// TIA Portal project "Parsing_migrated" (V16) (continued)
TYPE "LKinLang_typeKeyToken"
   STRUCT
      tokenBool : String["LKINLANG_LENGTH_OF_TOKEN_STRING"] := 'BOOL';   // Keyword for dataType "BOOL"
      tokenDInt : String["LKINLANG_LENGTH_OF_TOKEN_STRING"] := 'DINT';   // Keyword for dataType "DINT"
      tokenLReal : String["LKINLANG_LENGTH_OF_TOKEN_STRING"] := 'LREAL';   // Keyword for dataType "LREAL"
      tokenInterfaceVarBool : String["LKINLANG_LENGTH_OF_TOKEN_STRING"] := '%B';   // Keyword for interface variable type "BOOL"
      tokenInterfaceVarDInt : String["LKINLANG_LENGTH_OF_TOKEN_STRING"] := '%DI';   // Keyword for interface variable type "DINT"
      tokenInterfaceVarLReal : String["LKINLANG_LENGTH_OF_TOKEN_STRING"] := '%LR';   // Keyword for interface variable type "LREAL"
      tokenJumpTarget : String["LKINLANG_LENGTH_OF_TOKEN_STRING"] := 'LABEL';   // Keyword for label definition
      tokenJump : String["LKINLANG_LENGTH_OF_TOKEN_STRING"] := 'GOTO';   // Keyword for unconditional jump
      tokenJumpConditional : String["LKINLANG_LENGTH_OF_TOKEN_STRING"] := 'GOTOC';   // Keyword for conditional jump
      tokenPreprocessingStop : String["LKINLANG_LENGTH_OF_TOKEN_STRING"] := 'STOPRE';   // Keyword for preprocessing stop
      tokenIf : String["LKINLANG_LENGTH_OF_TOKEN_STRING"] := 'IF';   // Keyword for start of IF
      tokenElse : String["LKINLANG_LENGTH_OF_TOKEN_STRING"] := 'ELSE';   // Keyword for ELSE / Keyword for Else
      tokenEndIf : String["LKINLANG_LENGTH_OF_TOKEN_STRING"] := 'ENDIF';   // Keyword for end of IF / Keyword for end of if
      tokenWhile : String["LKINLANG_LENGTH_OF_TOKEN_STRING"] := 'WHILE';   // Keyword for start of WHILE
      tokenEndWhile : String["LKINLANG_LENGTH_OF_TOKEN_STRING"] := 'ENDWHILE';   // Keyword for end of WHILE
      tokenFor : String["LKINLANG_LENGTH_OF_TOKEN_STRING"] := 'FOR';   // Keyword for start of FOR
      tokenQuantity : String["LKINLANG_LENGTH_OF_TOKEN_STRING"] := 'TO';   // Keyword for end value of FOR
      tokenIncrement : String["LKINLANG_LENGTH_OF_TOKEN_STRING"] := 'STEP';   // Keyword for increment of FOR
      tokenEndFor : String["LKINLANG_LENGTH_OF_TOKEN_STRING"] := 'ENDFOR';   // Keyword for end of FOR
      tokenStartSub : String["LKINLANG_LENGTH_OF_TOKEN_STRING"] := 'SUB';   // Keyword for starting the definition of a subprogram
      tokenEndSub : String["LKINLANG_LENGTH_OF_TOKEN_STRING"] := 'ENDSUB';   // Keyword for ending the definition of a subprogram
      tokenCallSub : String["LKINLANG_LENGTH_OF_TOKEN_STRING"] := 'CALL';   // Keyword for calling a subprogram
      tokenReturnSub : String["LKINLANG_LENGTH_OF_TOKEN_STRING"] := 'RETURN';   // Keyword for returning from a subprogram
   END_STRUCT;
END_TYPE

TYPE "LKinLang_typeFlagModeDefaults"
   STRUCT
      setFlags : Array[0.."LKINCTRL_NO_OF_LAST_SETFLAG"] of "LKinLang_typeFlagModeDefaultElement";   // Default flag settings for respective setFlag number
      valueFlags : Array[0.."LKINCTRL_NO_OF_LAST_VALUEFLAG"] of "LKinLang_typeFlagModeDefaultElement";   // Default flag settings for respective valueFlag number
   END_STRUCT;
END_TYPE

TYPE "LKinLang_typeLineTokens"
   STRUCT
      lineNo : UDInt;   // line number
      numberOfToken : DInt;   // number of token
      lineToken : Array[1.."LKINLANG_MAX_NUMBER_OF_TOKEN_PER_LINE"] of String["LKINLANG_LENGTH_OF_TOKEN_STRING"];   // array of line tokens
   END_STRUCT;
END_TYPE

TYPE "LKinLang_typeMathParserResult"
   STRUCT
      finalResult : LReal;   // final result of math parser
      errorID : DInt;   // error code of math parser calculation
   END_STRUCT;
END_TYPE

TYPE "LKinLang_typeDiffElementaryDatatypes"
   STRUCT
      valueLReal : LReal;   // LReal value
      valueReal : Real;   // Real value
      valueDint : DInt;   // DInt value
      valueInt : Int;   // Int value
   END_STRUCT;
END_TYPE

TYPE "LKinLang_typeFlagModeDefaultElement"
   STRUCT
      flagMode : USInt;   // Default flag mode for respective setFlag number
      remainingDistance : LReal;   // Default remainingDistance for respective setFlag number in case of flagMode = 10
   END_STRUCT;
END_TYPE

TYPE "LKinLang_typePreProcessorReplacement"
   STRUCT
      replacements : Array[1.."LKINLANG_NUMBER_OF_REPLACEMENTS"] of Struct   // pre-processor replacement structure
         searchTerm : String["LKINLANG_MAX_NUMBER_OF_TOKEN_PER_LINE"];   // term to be searched
         replaceTerm : String["LKINLANG_MAX_NUMBER_OF_TOKEN_PER_LINE"];   // term to replace search term
      END_STRUCT;
   END_STRUCT;
END_TYPE

TYPE "LKinLang_typeGCodeDefaults"
   STRUCT
      velocityRapidLinear : LReal := -1.0;   // velocity for G0 command / velocity for FastLin command
      transitionVelocityMode : DInt := 5;   // Set G641 transition velocity (bufferMode); 2: low velocity, 5: high velocity
      orientationDirection : DInt := 3;   // Set orientation direction; 1: positive direction; 2: negative direction; 3: shortest distance
   END_STRUCT;
END_TYPE

TYPE "LKInLang_typeStackElement"
   STRUCT
      "type" : Int;   // Type of stack entry
      lineNumberStart : UDInt;   // Line number where stack entry starts
      lineNumberEnd : UDInt;   // Line number where stack entry ends
      variableRef : "LKinLang_typeVarRef";   // Counter variable reference (only for FOR loops)
      increment : DInt;   // Increment of FOR loop
      quantity : DInt;   // End value of FOR loop
   END_STRUCT;
END_TYPE

TYPE "LKInLang_typeHierarchicLevel"
   STRUCT
      currentLevel : Int;   // Current hierarchic level
      numberOfLevels : Int;   // Number of found hierarchic level changes
      levels : Array[1.."LKINLANG_NUMBER_OF_HIERARCHICLEVEL"] of "LKInLang_typeHierarchicLevelElement";   // Array of level changes
   END_STRUCT;
END_TYPE

TYPE "LKinLang_typeStack"
   STRUCT
      numberOfElements : Int;   // Counter for stack elements
      stackElements : Array[1..20] of "LKInLang_typeStackElement";   // Array of stack entries
   END_STRUCT;
END_TYPE

TYPE "LKInLang_typeHierarchicLevelElement"
   STRUCT
      lineNumber : UDInt;   // Line number where new hierarchic level start
      level : Int;   // Value of hierarchic level
      "type" : Int;   // Type of hierarchic level
   END_STRUCT;
END_TYPE

TYPE "LKinLang_typeSubPrg"
   STRUCT
      prgName : String;   // Name of subprogram
      lineNumberStart : UDInt;   // Line number where subprograms starts
      lineNumberEnd : UDInt;   // Line number where subprograms ends
   END_STRUCT;
END_TYPE

TYPE "LKinLang_typeSubPrgList"
   STRUCT
      numberOfSubPrgs : Int;   // Counter of found subprograms
      subPrgs : Array[1.."LKINLANG_NUMBER_OF_SUBPROGRAMS"] of "LKinLang_typeSubPrg";   // Array of subprograms
   END_STRUCT;
END_TYPE

TYPE "LKinLang_typeVariableDeclaration"
   STRUCT
      localVariables : String := 'DEF _type_ _name_';   // How to declare a local variable
      globalVariables : String := 'DEF GLOBAL _type_ _name_';   // How to declare a global variable
   END_STRUCT;
END_TYPE

TYPE "LKinLang_typeParameterDefinition"
   STRUCT
      parameterNameString : String;   // parameter name (textual)
      parameterNameNumber : DInt := -1;   // parameter name (numerical)
      properties : DWord;   // parameter properties
      validCountPerLine : Int := 1;   // counter of valid parameter uses per line
      directValues : "LKinCtrl_typePathDataElement_advanced";   // direct values in PathData element
      followingValues : Array[1.."LKINLANG_NUMBER_OF_FOLLOW_VALUES"] of "LKinLang_typePathDataBoolean";   // following values in PathData element variables (Boolean)
      priorities : "LKinLang_typePathDataElementCounter";   // priorities of PathData element variables (Int)
      conditions : Array[1.."LKINLANG_NUMBER_OF_CONDITIONS"] of "LKinLang_typeCondition";   // array of conditons
   END_STRUCT;
END_TYPE

TYPE "LKinLang_typePathDataElement"
   STRUCT
      pathDataElement : "LKinCtrl_typePathDataElement_advanced";   // PathData element
      priority : "LKinLang_typePathDataElementInteger";   // PathData element priorities (Int)
      properties : DWord;   // properties
      motionCmd : Int;   // number of motion command
   END_STRUCT;
END_TYPE

TYPE "LKinLang_typeCondition"
   STRUCT
      ParameterNumber : DInt;   // assignment to specific command
      Group : DInt;   // summarization of conditions
      Mode : DInt;   // specification where to evaulate conditions
   END_STRUCT;
END_TYPE

TYPE "LKinLang_typeLineContent"
   STRUCT
      number : UDInt;   // line number
      content : String["LKINLANG_LENGTH_OF_ASCII_LINE_STRING"];   // line content (textual)
   END_STRUCT;
END_TYPE

TYPE "LKinLang_typeLineBuffer"
   STRUCT
      info : "LKinLang_typeFileInfo";   // status of current loaded file
      pointers : "LKinLang_typeLineBufferPointer";   // pathData pointer structure / PathData pointer structure
      lines : Array["LKINLANG_FIRST_INDEX_LINE_BUFFER".."LKINLANG_LAST_INDEX_LINE_BUFFER"] of "LKinLang_typeLineContent";   // line buffer structure
   END_STRUCT;
END_TYPE

TYPE "LKinLang_typeParameterCounter"
   STRUCT
      parameterNumber : Int;   // number of paramter
      counterValue : Int;   // counter value
   END_STRUCT;
END_TYPE

TYPE "LKinLang_typeParameterLookUp"
   STRUCT
      parameterNameString : String;   // parameter name (textual)
      parameterNameNumber : DInt;   // parameter name (numerical)
      parameterNumber : Int;   // parameter number
      directValueWord : Word;   // direct value word
      followValueWords : Array[1.."LKINLANG_NUMBER_OF_FOLLOW_VALUES"] of Word;   // array of follow value words
   END_STRUCT;
END_TYPE

// folder: LKinLang_Types/LKinLang_typesBoolean

TYPE "LKinLang_typePathDataValid"
   STRUCT
      cmdType : Bool := FALSE;   // TRUE: Take FollowingValue as cmdType
      cmdName : Bool := FALSE;   // TRUE: Take FollowingValue as cmdName
      cmdCoordinates : "LKinLang_typeCoordsBoolean";   // Command coordinates
      cmdParameters : "LKinLang_typeParameterBoolean";   // Command parameters
      setFlags : Array[1.."LKINCTRL_NO_OF_CMD_SETFLAGS"] of "LKinLang_typeFlagBoolean";   // Flags to control actuators
      valueFlags : Array[1.."LKINCTRL_NO_OF_CMD_VALUEFLAGS"] of "LKinLang_typeValueFlagBoolean";   // Flags to control actuators
   END_STRUCT;
END_TYPE

TYPE "LKinLang_typeValueFlagBoolean"
   STRUCT
      flag : Bool;   // TRUE: Take FollowingValue as Flag
      value : Bool;
      flagMode : Bool;   // TRUE: Take FollowingValue as FlagMode
      remainingDistance : Bool;   // TRUE: Take FollowingValue as RemainingDistance
   END_STRUCT;
END_TYPE

TYPE "LKinLang_typeCoordsBoolean"
   STRUCT
      cartesianPosition : "LKinLang_typeCartPosBoolean";   // Cartesian position
      coordSystem : Bool;   // TRUE: Take FollowingValue as CoordSystem
   END_STRUCT;
END_TYPE

TYPE "LKinLang_typeCartPosBoolean"
   STRUCT
      x : Bool;   // TRUE: Take FollowingValue as X Position
      y : Bool;   // TRUE: Take FollowingValue as Y Position
      z : Bool;   // TRUE: Take FollowingValue as Z Position
      "a" : Bool;   // TRUE: Take FollowingValue as A Position
   END_STRUCT;
END_TYPE

TYPE "LKinLang_typeParameterBoolean"
   STRUCT
      pathDynamics : "LKinLang_typeDynamicsBoolean";   // Dynamic settings
      orientationDirection : Bool;   // TRUE: Take FollowingValue as OrientationDirection
      bufferMode : Bool;   // TRUE: Take FollowingValue as bufferMode
      transitionParameters : Array[1..5] of Bool;   // Blending parameters
      dynamicAdaption : Bool;   // TRUE: Take FollowingValue as DynamicAdaption
      offsetParameters : "LKinLang_typeOffsetParametersBoolean";   // Offset parameter
      circleParameters : "LKinLang_typeCircleParameterBoolean";   // Circle parameter
   END_STRUCT;
   // // transitionParameters[1] : TRUE: Take FollowingValue as TransitionParameter[1]
   // // transitionParameters[2] : TRUE: Take FollowingValue as TransitionParameter[2]
   // // transitionParameters[3] : TRUE: Take FollowingValue as TransitionParameter[3]
   // // transitionParameters[4] : TRUE: Take FollowingValue as TransitionParameter[4]
   // // transitionParameters[5] : TRUE: Take FollowingValue as TransitionParameter[5]
END_TYPE

TYPE "LKinLang_typeDynamicsBoolean"
   STRUCT
      velocity : Bool;   // TRUE: Take FollowingValue as Velocity
      acceleration : Bool;   // TRUE: Take FollowingValue as Acceleration
      deceleration : Bool;   // TRUE: Take FollowingValue as Deceleration
      jerk : Bool;   // TRUE: Take FollowingValue as Jerk
   END_STRUCT;
END_TYPE

TYPE "LKinLang_typeCircleParameterBoolean"
   STRUCT
      circMode : Bool;   // TRUE: Take FollowingValue as CircMode
      auxPoint : Array[1..3] of Bool;   // Circle aux point
      pathChoice : Bool;   // TRUE: Take FollowingValue as PathChoice
      circlePlane : Bool;   // TRUE: Take FollowingValue as CirclePlane
      radius : Bool;   // TRUE: Take FollowingValue as CircleRadius
      arc : Bool;   // TRUE: Take FollowingValue as CircleArc
   END_STRUCT;
   // // auxPoint[1] : TRUE: Take FollowingValue as AuxPoint[1]
   // // auxPoint[2] : TRUE: Take FollowingValue as AuxPoint[2]
   // // auxPoint[3] : TRUE: Take FollowingValue as AuxPoint[3]
END_TYPE

TYPE "LKinLang_typePathDataBoolean"
   STRUCT
      cmdType : Bool := FALSE;   // TRUE: Take FollowingValue as cmdType
      cmdName : Bool := FALSE;   // TRUE: Take FollowingValue as cmdName
      cmdCoordinates : "LKinLang_typeCoordsBoolean";   // Command coordinates
      cmdParameters : "LKinLang_typeParameterBoolean";   // Command parameters
      setFlags : "LKinLang_typeFlagBoolean";   // Flags to control actuators
      valueFlags : "LKinLang_typeValueFlagBoolean";
   END_STRUCT;
END_TYPE

TYPE "LKinLang_typeFlagBoolean"
   STRUCT
      flag : Bool;   // TRUE: Take FollowingValue as Flag
      flagMode : Bool;   // TRUE: Take FollowingValue as FlagMode
      remainingDistance : Bool;   // TRUE: Take FollowingValue as RemainingDistance
   END_STRUCT;
END_TYPE

TYPE "LKinLang_typeOffsetParametersBoolean"
   STRUCT
      offsetParaNo : Bool;   // TRUE: Take FollowingValue as OffsetParamNo
      mainPathPlane : Bool;   // TRUE: Take FollowingValue as MainPathPlane
   END_STRUCT;
END_TYPE

// folder: LKinLang_Types/LKinLang_typesCounter

TYPE "LKinLang_typeValueFlagInteger"
   STRUCT
      flag : Int;   // flag (priority)
      value : Int;
      flagMode : Int;   // flag mode (priority)
      remainingDistance : Int;   // remaining distance (priority)
   END_STRUCT;
END_TYPE

TYPE "LKinLang_typeCoordsInteger"
   STRUCT
      cartesianPosition : "LKinLang_typeCartPosInteger";   // cartesian target coordinats (priority)
      coordSystem : Int;   // coordinate system (priority)
   END_STRUCT;
END_TYPE

TYPE "LKinLang_typeCartPosInteger"
   STRUCT
      x : Int;   // X (priority)
      y : Int;   // Y (priority)
      z : Int;   // Z (priority)
      "a" : Int;   // A (priority)
   END_STRUCT;
END_TYPE

TYPE "LKinLang_typeParameterInteger"
   STRUCT
      pathDynamics : "LKinLang_typeDynamicsInteger";   // dynamic settings (priority)
      orientationDirection : Int;   // orientation direction (priority)
      bufferMode : Int;   // bufferMode (priority)
      transitionParameters : Array[1..5] of Int;   // blending parameters
      dynamicAdaption : Int;   // dynamicAdaption (priority)
      offsetParameters : "LKinLang_typeOffsetParameters";   // offset parameter
      circleParameters : "LKinLang_typeCircleParameterInteger";   // parameters for MoveCircAbs and MoveCircRel
   END_STRUCT;
END_TYPE

TYPE "LKinLang_typeDynamicsInteger"
   STRUCT
      velocity : Int;   // velocity (priority)
      acceleration : Int;   // acceleration (priority)
      deceleration : Int;   // deceleration (priority)
      jerk : Int;   // jerk (priority)
   END_STRUCT;
END_TYPE

TYPE "LKinLang_typeCircleParameterInteger"
   STRUCT
      circMode : Int;   // circMode (priority)
      auxPoint : Array[1..3] of Int;   // auxPoint (priority)
      endPoint : Array[1..4] of Int;   // endPoint (priority)
      pathChoice : Int;   // path choice (priority)
      circlePlane : Int;   // cicle Plane (priority)
      radius : Int;   // raduis (priority)
      arc : Int;   // arc (priority)
   END_STRUCT;
   // // auxPoint[1] : X (priority)
   // // auxPoint[2] : Y (priority)
   // // auxPoint[3] : Z (priority)
   // // endPoint[1] : X (priority)
   // // endPoint[2] : Y (priority)
   // // endPoint[3] : Z (priority)
   // // endPoint[4] : A (priority)
END_TYPE

TYPE "LKinLang_typePathDataElementInteger"
   STRUCT
      cmdType : Int := 0;   // 1: MoveLinAbs; 2: MoveLinRel; 3: MoveCircAbs; 4: MoveCircRel; -1: End of List
      cmdName : Int;   // name of command
      cmdCoordinates : "LKinLang_typeCoordsInteger";   // target coordinate definition (priority)
      cmdParameters : "LKinLang_typeParameterInteger";   // additional command parameters (priority)
      setFlags : Array[1.."LKINCTRL_NO_OF_CMD_SETFLAGS"] of "LKinLang_typeFlagInteger";   // setFlags (priority)
      valueFlags : Array[1.."LKINCTRL_NO_OF_CMD_VALUEFLAGS"] of "LKinLang_typeValueFlagInteger";   // setFlags (priority)
   END_STRUCT;
   // // cmdParameters.pathDynamics.velocity : velocity (priority)
   // // cmdParameters.pathDynamics.acceleration : acceleration (priority)
   // // cmdParameters.pathDynamics.deceleration : deceleration (priority)
   // // cmdParameters.pathDynamics.jerk : jerk (priority)
   // // cmdParameters.orientationDirection : orientation direction (priority)
   // // cmdParameters.bufferMode : bufferMode (priority)
   // // cmdParameters.transitionParameters : blending parameters (priority)
END_TYPE

TYPE "LKinLang_typePathDataElementCounter"
   STRUCT
      cmdType : Int := 0;   // 1: MoveLinAbs; 2: MoveLinRel; 3: MoveCircAbs; 4: MoveCircRel; -1: End of List
      cmdName : Int;   // name of command
      cmdCoordinates : "LKinLang_typeCoordsInteger";   // target coordinate definition
      cmdParameters : "LKinLang_typeParameterInteger";   // additional command parameters
      setFlags : "LKinLang_typeFlagInteger";   // flags to control actuators
      valueFlags : "LKinLang_typeValueFlagInteger";   // flags to control actuators
   END_STRUCT;
   // // cmdCoordinates.cartesianPosition : cartesian target coordinats
   // // cmdCoordinates.cartesianPosition.x : X
   // // cmdCoordinates.cartesianPosition.y : Y
   // // cmdCoordinates.cartesianPosition.z : Z
   // // cmdCoordinates.cartesianPosition."a" : A
   // // cmdCoordinates.coordSystem : 0: WCS; 1: OCS[1]; 2: OCS[2]; 3: OCS[3]
   // // cmdParameters.pathDynamics : dynamic settings
   // // cmdParameters.pathDynamics.velocity : >0.0: configured value used; <0.0: default TO setting used; for cmdType = 100 ==> waitTime in ms
   // // cmdParameters.pathDynamics.acceleration : >0.0: configured value used; <0.0: default TO setting used
   // // cmdParameters.pathDynamics.deceleration : >0.0: configured value used; <0.0: default TO setting used
   // // cmdParameters.pathDynamics.jerk : >0.0: configured value used; <0.0: default TO setting used
   // // cmdParameters.orientationDirection : 1: positive direction; 2: negative direction; 3: shortest distance
   // // cmdParameters.bufferMode : 1: standstill between commands, 2: blending with lower speed; 5: blending with higher speed
   // // cmdParameters.transitionParameters : blending parameters
   // // cmdParameters.transitionParameters[1] : blending distance - >0.0: configured value used; <0.0: maximum possible blending distance used
   // // cmdParameters.transitionParameters[2] : reserved, do not set
   // // cmdParameters.transitionParameters[3] : reserved, do not set
   // // cmdParameters.transitionParameters[4] : reserved, do not set
   // // cmdParameters.transitionParameters[5] : reserved, do not set
   // // cmdParameters.dynamicAdaption : <0.0: default TO setting used; 0: no dynamic adaption; 1: with variable limits; 2: with constant limits
   // // cmdParameters.offsetParameters : parameters for offset selection and configuration
   // // cmdParameters.offsetParameters.offsetParaNo : selection of offset parameter set from configuration structure
   // // cmdParameters.offsetParameters.mainPathPlane : main path plane for compensation
   // // cmdParameters.circleParameters : parameters for MoveCircAbs and MoveCircRel
   // // cmdParameters.circleParameters.circMode : 0: auxPoint defines point on circle line; 1: auxPoint defines circle center; 2: radius and endPoint define circle segment; 3: GCode notation (end & aux point)
   // // cmdParameters.circleParameters.auxPoint : auxiliary point for circle definition
   // // cmdParameters.circleParameters.auxPoint[1] : X
   // // cmdParameters.circleParameters.auxPoint[2] : Y
   // // cmdParameters.circleParameters.auxPoint[3] : Z
   // // cmdParameters.circleParameters.arc : only in combination with circMode(1): arc
   // // cmdParameters.circleParameters.radius : only in combination with circMode(2): radius
   // // cmdParameters.circleParameters.circlePlane : circMode(0): not relevant; circMode(1+2): 0: XZ; 1: YZ; 2: XY
   // // cmdParameters.circleParameters.pathChoice : circMode(0): not relevant; circMode(1): 0: pos direction; 1: neg direction; circMode(2): 0: short pos segment; 1: short neg segment; 2: long pos segment; 3: long neg segment
END_TYPE

TYPE "LKinLang_typeFlagInteger"
   STRUCT
      flag : Int;   // flag (priority)
      flagMode : Int;   // flag mode (priority)
      remainingDistance : Int;   // remaining distance (priority)
   END_STRUCT;
END_TYPE

TYPE "LKinLang_typeOffsetParameters"
   STRUCT
      offsetParaNo : Int;   // selection of offset parameter set from configuration structure
      mainPathPlane : Int;   // main path plane for compensation
   END_STRUCT;
END_TYPE

// folder: (top level)

DATA_BLOCK "DB_Writing"   // DB5
{ S7_Optimized_Access := 'TRUE' }
VERSION : 0.1
   VAR
      EnableAxes : Bool := false;   // control variable to enable axes with MC_POWER
      AxesEnabled : Bool := false;   // status variable to see all axes enabled
      ResetAxes : Bool := false;   // control variable to reset axes with MC_RESET
      AxesError : Bool := false;   // status variable to see error on one axis
      HomeAxes : Bool := false;   // control variable to home axes with MC_HOME
      AxesHomed : Bool := false;   // status variable to see all axes homed
      HomePos : Array[1..4] of LReal;   // control variable storing homing positions for MC_GroupHome
      HomeMode : Array[1..4] of Int;   // control variable storing homing modes for MC_GroupHome
      RestartMode : Array[1..5] of Bool;   // control variable storing restart modes for MC_GroupReset
      StartMode : Array[1..4] of DInt;   // control variable storing start modes for MC_GroupPower
      StopMode : Array[1..4] of Int;   // control variable storing stop modes for MC_GroupPower
      executeProgram : Bool := false;   // control variable to execute a program once
      stopProgram : Bool := false;   // control variable to stop the program execution
      resetProgram : Bool := false;
      textInput : String := '';
      textLength : DInt := 0;
   END_VAR
   VAR RETAIN
      maxTextLength : Int := 20;
      enterLenght : Int := 8;
   END_VAR
   VAR
      TextCharArray : Array[0..19] of Char;
   END_VAR
   VAR RETAIN
      beginPosFileName : String := 'gotobeginpos.nc';
      endPosFileName : String := 'gotohomepos.nc';
      fileNameCapsTemp : String := 'caps_';
      fileNameTemp : String := 'lowercase_';
      spaceString : String := ' ';
   END_VAR
   VAR
      filename : String := '';
      programStatusString : String := ' ';
      gcodeFileNames : Array[0..24] of String;
      gcodeFileNames_copy : Array[0..24] of String;
      programLength : Int := 0;
      triggerTextbox : Bool := false;
      oldTriggerTextbox : Bool := false;
      oldTriggerExecuteProgram : Bool := false;
      loadFile : Bool := false;   // control variable to execute FileHandler load file
      saveFile : Bool := false;   // control variable to execute FileHandler save file
      fileHandler_stop : Bool := false;   // control variable to stop FileHandler
      fileHandler_done : Bool := false;
      fileHandler_error : Bool := false;
      parser_execute : Bool := false;   // control variable to execute Parser
      parser_stop : Bool := false;   // control variable to stop Parser
      parser_done : Bool := false;
      parser_error : Bool := false;
      movePath_active : Bool := false;
      movePath_execute : Bool := false;
      movePath_reset : Bool := false;
      movePath_stop : Bool := false;
      movePath_status : Word := 16#0;
      movePath_interrupt : Bool := false;
      movePath_error : Bool := false;
      movePath_done : Bool := false;
      statActualStep : Int := 10;
      lineBuffer : "LKinLang_typeLineBuffer";   // LineBuffer structure
      pathData : "LKinCtrl_typePathData_advanced";   // PathData structure
      preProcessorConfig : "LKinLang_typePreProcessorReplacement";   // Preprocessor config to search & replace
      parameterDefaults : "LKinLang_typeGCodeDefaults";   // Default values for GCode commands
      flagModeDefaults : "LKinLang_typeFlagModeDefaults";   // Default values for flags
      interfaceVariables : "LKinLang_typeInterfaceVariables";   // Interface variables
      movePathConfiguration : "LKinCtrl_typeConfiguration";   // Configuration for MovePath
      booleanFlagArray : Array[0.."LKINCTRL_NO_OF_LAST_SETFLAG"] of Bool;   // Boolean flag array connected to MovePath
      valueFlagArray : Array[0.."LKINCTRL_NO_OF_LAST_VALUEFLAG"] of LReal;   // Value flag array connected to MovePath
      programDone : Bool;
   END_VAR
BEGIN
   HomePos[1] := 200.0;
   HomePos[2] := 200.0;
   HomePos[3] := 200.0;
   StartMode[1] := 1;
   StartMode[2] := 1;
   StartMode[3] := 1;
   StartMode[4] := 1;
END_DATA_BLOCK

// folder: Instances

DATA_BLOCK "LKinCtrl_MC_GroupPower_DB"   // DB6
{ S7_Optimized_Access := 'TRUE' }
AUTHOR : tech.team.motioncontrol@siemens.com
FAMILY : LKinCtrl
VERSION : 2.0
// stored: InstanceOfName LKinCtrl_MC_GroupPower
"LKinCtrl_MC_GroupPower"
BEGIN
END_DATA_BLOCK

DATA_BLOCK "LKinCtrl_MC_GroupReset_DB"   // DB7
{ S7_Optimized_Access := 'TRUE' }
AUTHOR : tech.team.motioncontrol@siemens.com
FAMILY : LKinCtrl
VERSION : 2.0
// stored: InstanceOfName LKinCtrl_MC_GroupReset
"LKinCtrl_MC_GroupReset"
BEGIN
END_DATA_BLOCK

DATA_BLOCK "LKinCtrl_MC_GroupHome_DB"   // DB8
{ S7_Optimized_Access := 'TRUE' }
AUTHOR : tech.team.motioncontrol@siemens.com
FAMILY : LKinCtrl
VERSION : 2.0
// stored: InstanceOfName LKinCtrl_MC_GroupHome
"LKinCtrl_MC_GroupHome"
BEGIN
END_DATA_BLOCK

DATA_BLOCK "LKinLang_Filehandler_DB"   // DB9
{ S7_Optimized_Access := 'TRUE' }
AUTHOR : tech.team.motioncontrol@siemens.com
FAMILY : LKinLang
VERSION : 1.1
// stored: InstanceOfName LKinLang_Filehandler
"LKinLang_Filehandler"
BEGIN
END_DATA_BLOCK

DATA_BLOCK "LKinLang_Parser_DB"   // DB10
{ S7_Optimized_Access := 'TRUE' }
AUTHOR : tech.team.motioncontrol@siemens.com
FAMILY : LKinLang
VERSION : 1.3
// stored: InstanceOfName LKinLang_Parser
"LKinLang_Parser"
BEGIN
END_DATA_BLOCK

DATA_BLOCK "LKinCtrl_MC_MovePath_DB"   // DB11
{ S7_Optimized_Access := 'TRUE' }
AUTHOR : tech.team.motioncontrol@siemens.com
FAMILY : LKinCtrl
VERSION : 3.0
// stored: InstanceOfName LKinCtrl_MC_MovePath
"LKinCtrl_MC_MovePath"
BEGIN
END_DATA_BLOCK

// folder: (top level)

DATA_BLOCK "PositioningAxis_Left"   // DB1, Motion_DB
{ S7_Optimized_Access := 'TRUE' }
AUTHOR : SIMATIC
FAMILY : MC_1500
VERSION : 5.0
// stored: InstanceOfName TO_PositioningAxis
"TO_PositioningAxis"
BEGIN
END_DATA_BLOCK

DATA_BLOCK "PositioningAxis_Right"   // DB2, Motion_DB
{ S7_Optimized_Access := 'TRUE' }
AUTHOR : SIMATIC
FAMILY : MC_1500
VERSION : 5.0
// stored: InstanceOfName TO_PositioningAxis
"TO_PositioningAxis"
BEGIN
END_DATA_BLOCK

DATA_BLOCK "PositioningAxis_3"   // DB3, Motion_DB
{ S7_Optimized_Access := 'TRUE' }
AUTHOR : SIMATIC
FAMILY : MC_1500
VERSION : 5.0
// stored: InstanceOfName TO_PositioningAxis
"TO_PositioningAxis"
BEGIN
END_DATA_BLOCK

DATA_BLOCK "Kinematics_1"   // DB4, Motion_DB
{ S7_Optimized_Access := 'TRUE' }
AUTHOR : SIMATIC
FAMILY : MC_1500
VERSION : 5.0
// stored: InstanceOfName TO_Kinematics
"TO_Kinematics"
BEGIN
END_DATA_BLOCK

FUNCTION "ProcessText" : Void   // FC1, LAD
{ S7_Optimized_Access := 'TRUE' }
VERSION : 0.1
   VAR_INPUT
      fileNameCapsTemp : String;
      fileNameTemp : String;
      beginPosFileName : String;
      endPosFileName : String;
      textInput : String;
      textCharArray : Array[0..19] of Char;
      spaceString : String;
   END_VAR
   VAR_OUTPUT
      gcodeFileNames : Array[0..24] of String;
      programLength : Int;
   END_VAR
   VAR_TEMP
      i : Int;
      cnt : Int;
      TempString : String;
      TempString2 : String;
      FileName : String;
      stringInAscii : Int;
      "counter" : Int;
      numberofenters : Int;
   END_VAR
BEGIN

REGION Network 1 (SCL): Construction of the array of commands, select the right g code files
   // Go to begin position first before writing (letters are defined relative to begin position)
   "DB_Writing".gcodeFileNames[0] := #beginPosFileName;

   // Convert input string to array of chars
   Strg_TO_Chars(Strg := #textInput,
                 pChars := 0,
                 Cnt => "DB_Writing".textLength,
                 Chars := #textCharArray);

   // Loop over array of chars, make the file names
   #counter := 0;
   #numberofenters := 0;
   FOR #i := 1 TO "DB_Writing".textLength BY 1 DO
       #counter := #counter + 1;

       Chars_TO_Strg(Chars := #textCharArray,
                     pChars := #i - 1,
                     Cnt := 1,
                     Strg => #TempString);
       #stringInAscii := #textCharArray[#i - 1];

       // Ascii value between 65 and 90 --> uppercase letter
       IF (#stringInAscii >= 65 AND #stringInAscii <= 90) THEN
           #TempString2 := CONCAT(IN1 := #fileNameCapsTemp, IN2 := #TempString);

       // Not uppercase
       ELSE

           // A space is detected
           IF (#TempString = #spaceString) THEN
               #TempString2 := 'space';

           // Lowercase
           ELSE
               #TempString2 := CONCAT(IN1 := #fileNameTemp, IN2 := #TempString);
           END_IF;

       END_IF;

       #FileName := CONCAT(IN1 := #TempString2, IN2 := '.nc');
       "DB_Writing".gcodeFileNames[#counter] := #FileName;

       // An enter is detected or the text is going out of bounds
       IF (#stringInAscii = 10) OR (#i MOD "DB_Writing".enterLenght = 0) AND NOT (#i = "DB_Writing".textLength) THEN
           #counter := #counter + 1;
           "DB_Writing".gcodeFileNames[#counter] := 'enter.nc';
           #numberofenters := #numberofenters + 1;
       END_IF;

   END_FOR;

   // Go to end position
   #programLength := "DB_Writing".textLength + 2 + #numberofenters;
   "DB_Writing".gcodeFileNames[#programLength - 1] := #endPosFileName;

   // Reset rest of array
   FOR #i := #programLength TO "DB_Writing".maxTextLength + 1 + #numberofenters BY 1 DO
       "DB_Writing".gcodeFileNames[#i] := '';
   END_FOR;

   // Give as output
   #gcodeFileNames := "DB_Writing".gcodeFileNames;

   // Make a copy, because other array will be processed
   "DB_Writing".gcodeFileNames_copy := #gcodeFileNames;
END_REGION
END_FUNCTION

FUNCTION "Write" : Void   // FC2, LAD
{ S7_Optimized_Access := 'TRUE' }
VERSION : 0.1
   VAR_TEMP
      i : Int;
      dummyArray : Array[0..24] of String;
   END_VAR
BEGIN

REGION Network 1 (SCL): Loading/parsing/writing, main loop of program
   // Idea 1: write strings to know where we are in program, display on HMI - done
   // Idea 2: give error messages to HMI and display them
   "DB_Writing".filename := "DB_Writing".gcodeFileNames[0];

   IF LEN("DB_Writing".filename) > 0 THEN

       CASE "DB_Writing".statActualStep OF

           10: // Load NC file from memory
               "DB_Writing".loadFile := TRUE;
               "DB_Writing".programStatusString := CONCAT(IN1 := 'Loading ', IN2 := "DB_Writing".filename);

               IF "DB_Writing".fileHandler_done AND NOT "DB_Writing".fileHandler_error THEN
                   "DB_Writing".statActualStep := 20;
                   "DB_Writing".loadFile := FALSE;
               END_IF;

           20: // Parse NC file 
               "DB_Writing".parser_execute := TRUE;
               "DB_Writing".programStatusString := CONCAT(IN1 := 'Parsing ', IN2 := "DB_Writing".filename);

               IF "DB_Writing".parser_done AND NOT "DB_Writing".parser_error THEN
                   "DB_Writing".statActualStep := 30;
                   "DB_Writing".parser_execute := FALSE;
               END_IF;

           30: // Move
               "DB_Writing".movePath_execute := TRUE;
               "DB_Writing".programStatusString := CONCAT(IN1 := 'Writing ', IN2 := "DB_Writing".filename);

               IF "DB_Writing".movePath_done AND NOT "DB_Writing".movePath_error THEN
                   "DB_Writing".statActualStep := 40;
                   "DB_Writing".movePath_execute := FALSE;
               END_IF;

           40: // Initiate new array, shifted by one place, delete first entry of previous array
               "DB_Writing".programStatusString := 'Making array';

               FOR #i := 1 TO "DB_Writing".programLength - 1 DO
                   #dummyArray[#i - 1] := "DB_Writing".gcodeFileNames[#i];
               END_FOR;

               #dummyArray["DB_Writing".programLength - 1] := '';
               "DB_Writing".gcodeFileNames := #dummyArray;
               "DB_Writing".statActualStep := 10;

       END_CASE;

   ELSE
       "DB_Writing".programStatusString := 'Program finished';
       "DB_Writing".programDone := TRUE;
   END_IF;
END_REGION

REGION Network 2: Call LKinLang_FileHandler - read file from card
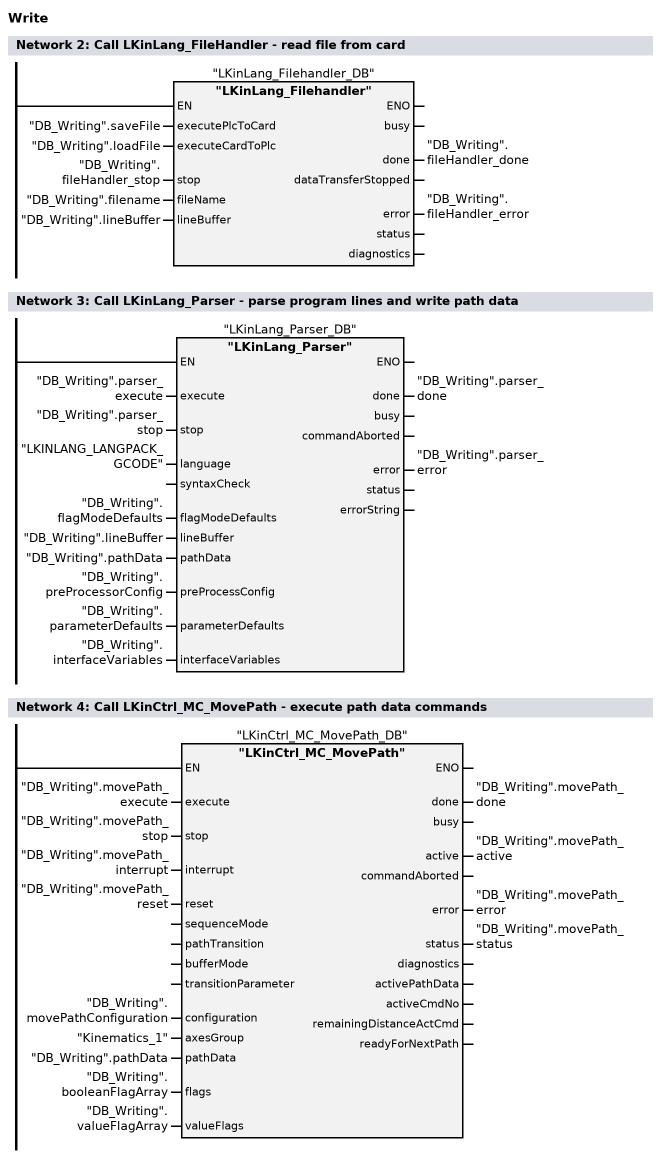
   RUNG wire#powerrail
      "LKinLang_Filehandler_DB"(executePlcToCard := "DB_Writing".saveFile, executeCardToPlc := "DB_Writing".loadFile, stop := "DB_Writing".fileHandler_stop, fileName := "DB_Writing".filename, lineBuffer := "DB_Writing".lineBuffer, busy =>, done => "DB_Writing".fileHandler_done, dataTransferStopped =>, error => "DB_Writing".fileHandler_error, status =>, diagnostics =>)
   END_RUNG
   // the same network as SCL:
   "LKinLang_Filehandler_DB"(executePlcToCard := "DB_Writing".saveFile,   // "LKinLang_Filehandler"
                           executeCardToPlc := "DB_Writing".loadFile,
                           stop := "DB_Writing".fileHandler_stop,
                           fileName := "DB_Writing".filename,
                           lineBuffer := "DB_Writing".lineBuffer,
                           done => "DB_Writing".fileHandler_done,
                           error => "DB_Writing".fileHandler_error);
END_REGION

REGION Network 3: Call LKinLang_Parser - parse program lines and write path data
   RUNG wire#powerrail
      "LKinLang_Parser_DB"(execute := "DB_Writing".parser_execute, stop := "DB_Writing".parser_stop, language := "LKINLANG_LANGPACK_GCODE", syntaxCheck :=, flagModeDefaults := "DB_Writing".flagModeDefaults, lineBuffer := "DB_Writing".lineBuffer, pathData := "DB_Writing".pathData, preProcessConfig := "DB_Writing".preProcessorConfig, parameterDefaults := "DB_Writing".parameterDefaults, interfaceVariables := "DB_Writing".interfaceVariables, done => "DB_Writing".parser_done, busy =>, commandAborted =>, error => "DB_Writing".parser_error, status =>, errorString =>)
   END_RUNG
   // the same network as SCL:
   "LKinLang_Parser_DB"(execute := "DB_Writing".parser_execute,   // "LKinLang_Parser"
                        stop := "DB_Writing".parser_stop,
                        language := "LKINLANG_LANGPACK_GCODE",
                        flagModeDefaults := "DB_Writing".flagModeDefaults,
                        lineBuffer := "DB_Writing".lineBuffer,
                        pathData := "DB_Writing".pathData,
                        preProcessConfig := "DB_Writing".preProcessorConfig,
                        parameterDefaults := "DB_Writing".parameterDefaults,
                        interfaceVariables := "DB_Writing".interfaceVariables,
                        done => "DB_Writing".parser_done,
                        error => "DB_Writing".parser_error);
END_REGION

REGION Network 4: Call LKinCtrl_MC_MovePath - execute path data commands
   RUNG wire#powerrail
      "LKinCtrl_MC_MovePath_DB"(execute := "DB_Writing".movePath_execute, stop := "DB_Writing".movePath_stop, interrupt := "DB_Writing".movePath_interrupt, reset := "DB_Writing".movePath_reset, sequenceMode :=, pathTransition :=, bufferMode :=, transitionParameter :=, configuration := "DB_Writing".movePathConfiguration, axesGroup := "Kinematics_1", pathData := "DB_Writing".pathData, flags := "DB_Writing".booleanFlagArray, valueFlags := "DB_Writing".valueFlagArray, done => "DB_Writing".movePath_done, busy =>, active => "DB_Writing".movePath_active, commandAborted =>, error => "DB_Writing".movePath_error, status => "DB_Writing".movePath_status, diagnostics =>, activePathData =>, activeCmdNo =>, remainingDistanceActCmd =>, readyForNextPath =>)
   END_RUNG
   // the same network as SCL:
   "LKinCtrl_MC_MovePath_DB"(execute := "DB_Writing".movePath_execute,   // "LKinCtrl_MC_MovePath"
                           stop := "DB_Writing".movePath_stop,
                           interrupt := "DB_Writing".movePath_interrupt,
                           reset := "DB_Writing".movePath_reset,
                           configuration := "DB_Writing".movePathConfiguration,
                           axesGroup := "Kinematics_1",
                           pathData := "DB_Writing".pathData,
                           flags := "DB_Writing".booleanFlagArray,
                           valueFlags := "DB_Writing".valueFlagArray,
                           done => "DB_Writing".movePath_done,
                           active => "DB_Writing".movePath_active,
                           error => "DB_Writing".movePath_error,
                           status => "DB_Writing".movePath_status);
END_REGION
END_FUNCTION

ORGANIZATION_BLOCK "Main"   // OB1, LAD, ProgramCycle
TITLE = "Main Program Sweep (Cycle)"
{ S7_Optimized_Access := 'TRUE' }
VERSION : 0.1
// Basic Motion Control commands for TO_PositioningAxis and TO_Kinematics
   VAR_INPUT
      Initial_Call : Bool;   // Initial call of this OB
      Remanence : Bool;   // =True, if remanent data are available
   END_VAR
BEGIN

REGION Network 1: Call LKinCtrl_MC_GroupPower - enable all axes interconnected with TO_Kinematics
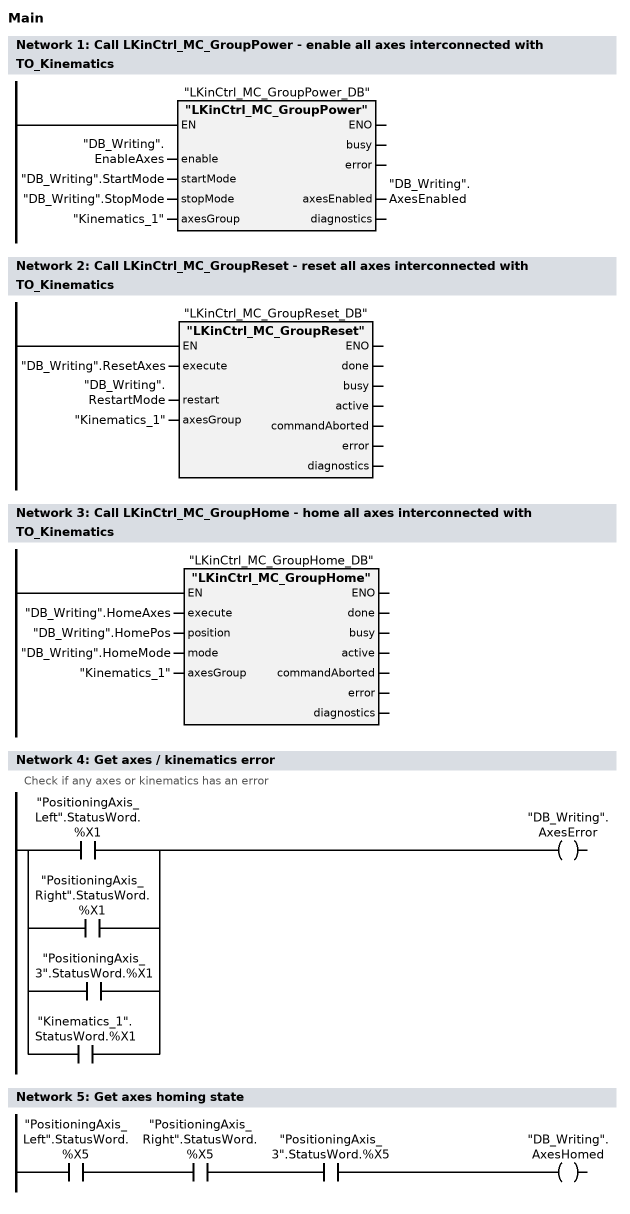
   RUNG wire#powerrail
      "LKinCtrl_MC_GroupPower_DB"(enable := "DB_Writing".EnableAxes, startMode := "DB_Writing".StartMode, stopMode := "DB_Writing".StopMode, axesGroup := "Kinematics_1", busy =>, error =>, axesEnabled => "DB_Writing".AxesEnabled, diagnostics =>)
   END_RUNG
   // the same network as SCL:
   "LKinCtrl_MC_GroupPower_DB"(enable := "DB_Writing".EnableAxes,   // "LKinCtrl_MC_GroupPower"
                           startMode := "DB_Writing".StartMode,
                           stopMode := "DB_Writing".StopMode,
                           axesGroup := "Kinematics_1",
                           axesEnabled => "DB_Writing".AxesEnabled);
END_REGION

REGION Network 2: Call LKinCtrl_MC_GroupReset - reset all axes interconnected with TO_Kinematics
   RUNG wire#powerrail
      "LKinCtrl_MC_GroupReset_DB"(execute := "DB_Writing".ResetAxes, restart := "DB_Writing".RestartMode, axesGroup := "Kinematics_1", done =>, busy =>, active =>, commandAborted =>, error =>, diagnostics =>)
   END_RUNG
   // the same network as SCL:
   "LKinCtrl_MC_GroupReset_DB"(execute := "DB_Writing".ResetAxes,   // "LKinCtrl_MC_GroupReset"
                           restart := "DB_Writing".RestartMode,
                           axesGroup := "Kinematics_1");
END_REGION

REGION Network 3: Call LKinCtrl_MC_GroupHome - home all axes interconnected with TO_Kinematics
   RUNG wire#powerrail
      "LKinCtrl_MC_GroupHome_DB"(execute := "DB_Writing".HomeAxes, position := "DB_Writing".HomePos, mode := "DB_Writing".HomeMode, axesGroup := "Kinematics_1", done =>, busy =>, active =>, commandAborted =>, error =>, diagnostics =>)
   END_RUNG
   // the same network as SCL:
   "LKinCtrl_MC_GroupHome_DB"(execute := "DB_Writing".HomeAxes,   // "LKinCtrl_MC_GroupHome"
                           position := "DB_Writing".HomePos,
                           mode := "DB_Writing".HomeMode,
                           axesGroup := "Kinematics_1");
END_REGION

REGION Network 4: Get axes / kinematics error
   // Check if any axes or kinematics has an error
   RUNG wire#powerrail
      Contact( "PositioningAxis_Left".StatusWord.%X1 )
      wire#w1
      Coil( "DB_Writing".AxesError )
   END_RUNG
   RUNG wire#powerrail
      Contact( "PositioningAxis_Right".StatusWord.%X1 )
   END_RUNG wire#w1
   RUNG wire#powerrail
      Contact( "PositioningAxis_3".StatusWord.%X1 )
   END_RUNG wire#w1
   RUNG wire#powerrail
      Contact( "Kinematics_1".StatusWord.%X1 )
   END_RUNG wire#w1
   // the same network as SCL:
   "DB_Writing".AxesError := "PositioningAxis_Left".StatusWord.%X1 OR "PositioningAxis_Right".StatusWord.%X1 OR "PositioningAxis_3".StatusWord.%X1 OR "Kinematics_1".StatusWord.%X1;
END_REGION

REGION Network 5: Get axes homing state
   RUNG wire#powerrail
      Contact( "PositioningAxis_Left".StatusWord.%X5 )
      Contact( "PositioningAxis_Right".StatusWord.%X5 )
      Contact( "PositioningAxis_3".StatusWord.%X5 )
      Coil( "DB_Writing".AxesHomed )
   END_RUNG
   // the same network as SCL:
   "DB_Writing".AxesHomed := "PositioningAxis_Left".StatusWord.%X5 AND "PositioningAxis_Right".StatusWord.%X5 AND "PositioningAxis_3".StatusWord.%X5;
END_REGION
END_ORGANIZATION_BLOCK

ORGANIZATION_BLOCK "WriteMain"   // OB123, LAD, ProgramCycle
TITLE = "Main Program Sweep (Cycle)"
{ S7_Optimized_Access := 'TRUE' }
VERSION : 0.1
   VAR_INPUT
      Initial_Call : Bool;   // Initial call of this OB
      Remanence : Bool;   // =True, if remanent data are available
   END_VAR
BEGIN

REGION Network 1 (SCL): Program logic to stop all FBs at once
   // Stop all FBs at once with "stopProgram"
   IF "DB_Writing".stopProgram THEN
       "DB_Writing".fileHandler_stop := TRUE;
       "DB_Writing".parser_stop := TRUE;
       "DB_Writing".movePath_stop := TRUE;
   END_IF;

   // Falling edge of stop program
   "FTrigStopProgram_DB"(CLK:="DB_Writing".stopProgram);

   // Reset stop bits when falling edge is detected
   IF "FTrigStopProgram_DB".Q THEN
       "DB_Writing".fileHandler_stop := FALSE;
       "DB_Writing".parser_stop := FALSE;
       "DB_Writing".movePath_stop := FALSE;
   END_IF;
END_REGION

REGION Network 2 (SCL): Program logic to reset axes and movePath FB at once
   // Reset all FBs at once with "resetProgram"
   IF "DB_Writing".resetProgram THEN
       "DB_Writing".movePath_reset := TRUE;
       "DB_Writing".ResetAxes := TRUE;
   END_IF;

   // Falling edge of reset program
   "FtrigResetProgram_DB"(CLK:="DB_Writing".resetProgram);

   // Reset stop bits when falling edge is detected
   IF "FtrigResetProgram_DB".Q THEN
       "DB_Writing".movePath_reset := FALSE;
       "DB_Writing".ResetAxes := FALSE;
   END_IF;
END_REGION

REGION Network 3 (SCL): Reset programDone bool on rising edge
   // Act when rising edge of trigger for processing text (set in HMI) is detected
   IF "DB_Writing".triggerTextbox AND NOT "DB_Writing".oldTriggerTextbox THEN
       "DB_Writing".programDone := FALSE;
   END_IF;

   "DB_Writing".oldTriggerTextbox := "DB_Writing".triggerTextbox;
END_REGION

REGION Network 4 (SCL): (Re-)initialize step value when pressing executeProgram/Get the letters from the input text block into array of readable file names on a rising edge
   // Act when rising edge of trigger executeProgram is detected
   IF "DB_Writing".executeProgram AND NOT "DB_Writing".oldTriggerExecuteProgram THEN
       "ProcessText"(fileNameCapsTemp := "DB_Writing".fileNameCapsTemp,
                     fileNameTemp := "DB_Writing".fileNameTemp,
                     beginPosFileName := "DB_Writing".beginPosFileName,
                     endPosFileName := "DB_Writing".endPosFileName,
                     textInput := "DB_Writing".textInput,
                     textCharArray := "DB_Writing".TextCharArray,
                     spaceString := "DB_Writing".spaceString,
                     gcodeFileNames => "DB_Writing".gcodeFileNames,
                     programLength => "DB_Writing".programLength);
       "DB_Writing".statActualStep := 10;
       "DB_Writing".gcodeFileNames := "DB_Writing".gcodeFileNames_copy; // reset the commands to an original copy
       "DB_Writing".programDone := FALSE;
   END_IF;

   "DB_Writing".oldTriggerExecuteProgram := "DB_Writing".executeProgram;
END_REGION

REGION Network 5: Enable write block
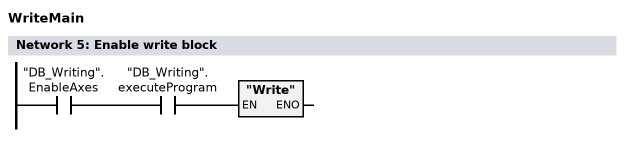
   RUNG wire#powerrail
      Contact( "DB_Writing".EnableAxes )
      Contact( "DB_Writing".executeProgram )
      "Write"()
   END_RUNG
   // the same network as SCL:
   IF "DB_Writing".EnableAxes AND "DB_Writing".executeProgram THEN "Write"(); END_IF;
END_REGION
END_ORGANIZATION_BLOCK

// folder: LKinCtrl_Blocks

